
               END_IF;
           END_REGION

       END_IF;
   END_REGION
END_FUNCTION

FUNCTION "Order State: Enter Requested Critical" : Void   // FC16, SCL
{ S7_Optimized_Access := 'TRUE' }
VERSION : 0.1
   VAR_INPUT
      timerVal : Real;
   END_VAR
   VAR_IN_OUT
      state : Int;
   END_VAR
   VAR_TEMP
      temp : Real;
   END_VAR
BEGIN
   IF #state = "requested" THEN
       IF #timerVal > 0.0 AND #timerVal <= "DEFAULT_CRITICAL_TIME" THEN
           #state := "requestedCrit";
       END_IF;
   END_IF;
END_FUNCTION

FUNCTION "Order State: Enter Requested Expired" : Void   // FC17, SCL
{ S7_Optimized_Access := 'TRUE' }
VERSION : 0.1
   VAR_INPUT
      timerVal : Real;
   END_VAR
   VAR_IN_OUT
      state : Int;
   END_VAR
BEGIN
   IF #state = "requestedCrit" THEN
       IF #timerVal <= -0.001 THEN
           #state := "requestedExp";
       END_IF;
   END_IF;
END_FUNCTION

// folder: Order/Timers

FUNCTION_BLOCK "Order Timer"   // FB6, SCL
{ S7_Optimized_Access := 'TRUE' }
VERSION : 0.1
   VAR_INPUT
      pnLib : "Recipe: PN Text Library";
   END_VAR
   VAR_IN_OUT
      stns : "Station: All Stations";
   END_VAR
   VAR
      rt : "Runtime Data";
   END_VAR
   VAR_TEMP
      pStn : Int;
      pBtn : Int;
   END_VAR
BEGIN
   REGION "RUNTIME CALL"
       #rt.elapsed := RUNTIME(#rt.mem);
       #rt.asReal := LREAL_TO_REAL(#rt.elapsed);
   END_REGION

   REGION "FOR EACH STATION"
       FOR #pStn := 0 TO "STATION_COUNT" DO

           REGION "FOR EACH BUTTON"
               FOR #pBtn := 0 TO "STATION_BUTTON_COUNT" DO

                   REGION "INITIALIZE TIMERS"
                       "Order Timer: Initialize"(pnLib := #pnLib,
                                                 pBtn := #pBtn,
                                                 stn := #stns.stn[#pStn]);
                   END_REGION

                   REGION "EXECUTE TIMERS"
                       "Order Timer: Timer Execution"(elapsedTime := #rt.asReal,
                                                      pBtn := #pBtn,
                                                      stn:=#stns.stn[#pStn],
                                                      timers := #stns.stn[#pStn].wipCmpts.timers);
                   END_REGION

               END_FOR;
           END_REGION

       END_FOR;
   END_REGION
END_FUNCTION_BLOCK

FUNCTION "Order Timer: Initialize" : Void   // FC8, SCL
{ S7_Optimized_Access := 'TRUE' }
VERSION : 0.1
   VAR_INPUT
      pnLib : "Recipe: PN Text Library";
      pBtn : Int;
   END_VAR
   VAR_IN_OUT
      stn : "Station: Single Station";
   END_VAR
   VAR_TEMP
      pnGood : Bool;
      default : Bool;
      clear : Bool;
   END_VAR
BEGIN
   REGION "ON PN CHANGE"
       IF #stn.wipCmpts.flags.newPN THEN

           REGION "INITIALIZE TO DEFAULT"

               REGION "EXECUTION VALIDATION"
                   #default := "Order Timer: Set to Default Check"(pnGood := #stn.wipCmpts.flags.pnGood[#pBtn],
                                                                   inSettingsScreen := #stn.wipCmpts.flags.inSettingsScreen,
                                                                   timerReset := #stn.wipCmpts.flags.resetTimer[#pBtn]);
               END_REGION

               REGION "ON VALIDATION"
                   IF #default THEN

                       REGION "SET DEFAULT TIME VALUE"
                           #stn.wipCmpts.timers.ptAllotted[#pBtn] := "DEFAULT_TOTAL_TIME";
                           #stn.wipCmpts.timers.ptCritical[#pBtn] := "DEFAULT_CRITICAL_TIME";
                       END_REGION

                   END_IF;
               END_REGION

           END_REGION

           REGION "INITIALIZE TO ZERO"

               REGION "EXECUTION VALIDATION"
                   #clear := "Order Timer: Set to Zero Check"(pnGood := #stn.wipCmpts.flags.pnGood[#pBtn],
                                                              inSettingsScreen := #stn.wipCmpts.flags.inSettingsScreen,
                                                              timerReset := #stn.wipCmpts.flags.resetTimer[#pBtn]);
               END_REGION

               REGION "ON VALIDATION"
                   IF #clear THEN

                       REGION "SET DEFAULT TIME VALUE"
                           #stn.wipCmpts.timers.ptAllotted[#pBtn] := 0.0;
                           #stn.wipCmpts.timers.ptCritical[#pBtn] := 0.0;
                       END_REGION

                   END_IF;
               END_REGION

           END_REGION

       END_IF;
   END_REGION
END_FUNCTION

FUNCTION "Order Timer: Timer Execution" : Void   // FC11, SCL
{ S7_Optimized_Access := 'TRUE' }
VERSION : 0.1
   VAR_INPUT
      elapsedTime : Real;
      pBtn : Int;
      stn : "Station: Single Station";
   END_VAR
   VAR_IN_OUT
      timers : "Station: Timers";
   END_VAR
BEGIN
   REGION "RUN CONDITIONS"
       CASE #stn.wipCmpts.orderState[#pBtn] OF

           "reset", "idle":
               IF #stn.flags.stateTransition[#pBtn] THEN
                   #timers.elapsed[#pBtn] := 0.0;
                   #timers.remaining[#pBtn] := 0.0;
               END_IF;

           "requested".."acknowledgedExp":
               #timers.elapsed[#pBtn] += #elapsedTime;
               #timers.remaining[#pBtn] := #timers.ptAllotted[#pBtn] - #timers.elapsed[#pBtn];

           ELSE:
               ;

       END_CASE;
   END_REGION
END_FUNCTION

FUNCTION "Order Timer: Set to Default Check" : Bool   // FC12, SCL
{ S7_Optimized_Access := 'TRUE' }
VERSION : 0.1
   VAR_INPUT
      pnGood : Bool;
      inSettingsScreen : Bool;
      timerReset : Bool;
   END_VAR
   VAR_TEMP
      ret : Bool;
   END_VAR
BEGIN
   REGION "ON VALID PN"
       #ret := #pnGood;
   END_REGION

   REGION "NOT WHILE IN SETTINGS SCREEN"
       IF #inSettingsScreen THEN
           #ret := FALSE;
       END_IF;
   END_REGION

   REGION "ON RESET REQUEST"
       #ret := #timerReset OR #ret;
   END_REGION

   REGION "RETURN"
       #"Order Timer: Set to Default Check" := #ret;
   END_REGION
END_FUNCTION

FUNCTION "Order Timer: Set to Zero Check" : Bool   // FC15, SCL
{ S7_Optimized_Access := 'TRUE' }
VERSION : 0.1
   VAR_INPUT
      pnGood : Bool;
      inSettingsScreen : Bool;
      timerReset : Bool;
   END_VAR
   VAR_TEMP
      ret : Bool;
   END_VAR
BEGIN
   REGION "ON VALID PN"
       #ret := NOT #pnGood;
   END_REGION

   REGION "NOT WHILE IN SETTINGS SCREEN"
       IF #inSettingsScreen THEN
           #ret := FALSE;
       END_IF;
   END_REGION

   REGION "ON RESET REQUEST"
       #ret := #timerReset OR #ret;
   END_REGION

   REGION "RETURN"
       #"Order Timer: Set to Zero Check" := #ret;
   END_REGION
END_FUNCTION

// folder: Part Request

FUNCTION_BLOCK "Part Request"   // FB7, SCL
{ S7_Optimized_Access := 'TRUE' }
VERSION : 0.1
   VAR_INPUT
      stns : "Station: All Stations";
      savedWips : "Recipe: HMI Stations Saved Wips";
      pnLib : "Recipe: PN Text Library";
   END_VAR
   VAR_IN_OUT
      dataTable : "Part Request Data";
   END_VAR
   VAR RETAIN
      pDataRow : Int;
   END_VAR
   VAR_TEMP
      address : DInt;
      addRequest : Bool;
      inTable : DInt;
      pStn : Int;
      pBtn : Int;
      pWip : Int;
      pRqstsRow : Int;
      removeRequest : Bool;
   END_VAR
BEGIN
   REGION "FOR EACH STATION"
       FOR #pStn := 0 TO "STATION_COUNT" DO

           REGION "FOR EACH BUTTON"
               FOR #pBtn := 0 TO "STATION_BUTTON_COUNT" DO

                   REGION "NEXT BUTTON ON NO TRANSITION"
                       IF NOT #stns.stn[#pStn].flags.stateTransition[#pBtn] THEN
                           GOTO NOSTNREQ;
                       END_IF;
                   END_REGION

                   REGION "GET ADDRESS"
                       #pWip := DINT_TO_INT(#stns.stn[#pStn].wipData.index);
                       #address := "Address.Set_Address"(pStn := #pStn, pBtn := #pBtn, pWip := #pWip);
                   END_REGION

                   REGION "CHECK FOR ENTRY IN DATA TABLE"
                       #inTable := "Part Request: Address in Table"(search := #address,
                                                                    dataTable := #dataTable);
                   END_REGION

                   REGION "ADD"

                       REGION "VALIDATE CONDITIONS"
                           #addRequest := "Part Request: Validate Add"(inTable := #inTable,
                                                                       orderState := #stns.stn[#pStn].wipCmpts.orderState[#pBtn]);
                       END_REGION

                       REGION "EXECUTE"
                           IF #addRequest THEN
                               #addRequest := FALSE;
                               #dataTable.row[#pDataRow] := #address;
                               "Row Pointer: Roll Over"(limit := "partReqDataRowCount",
                                                                "pointer" := #pDataRow);
                           END_IF;
                       END_REGION

                   END_REGION

                   REGION "REMOVE SINGLE STATION"

                       REGION "VALIDATE CONDITIONS: SINGLE"
                           #removeRequest := "Part Request: Validate Remove: Single"(inTable := #inTable,
                                                                                     orderState := #stns.stn[#pStn].wipCmpts.orderState[#pBtn]);
                       END_REGION

                       REGION "EXECUTE"
                           IF #removeRequest THEN
                               #removeRequest := FALSE;
                               #dataTable.row[#inTable] := -1;
                               "Part Request: Collapse Table"(#dataTable);
                               "Row Pointer: Post Collapse"(dataTable := #dataTable,
                                                            pDataRow := #pDataRow);
                           END_IF;
                       END_REGION

                   END_REGION

               NOSTNREQ:
                   ;
               END_FOR;
           END_REGION

       END_FOR;
   END_REGION


   (* REGION "REMOVE WIP STATIONS"                    
       FOR #pStn := 0 TO "hmiStnCount" DO
           FOR #pWip := 0 TO "wipCount" DO
               IF #savedWips.stn[#pStn].wip[#pWip].flags.clearWipRequest THEN
                   FOR #pBtn := 0 TO "btnCount" DO
                       #address := "Address: Set Address"(pBtn := #pBtn, pStn := #pStn, pWip := #pWip);
                       #inTable := "Part Request: Address in Table"(adrRequest := #address,
                                                                    dataTable := #dataTable);
                       #removeRequest := "Part Request: Validate Remove: WIP"(inTable := #inTable,
                                                                              clearWipRequest := #savedWips.stn[#pStn].wip[#pWip].flags.clearWipRequest);
                       IF #removeRequest THEN
                           #removeRequest := FALSE;
                           "Part Request: Remove"(pRow := #inTable,
                                                  dataTable := #dataTable);
                           "Part Request: Collapse Table"(#dataTable);
                           "Row Pointer: Post Collapse"(dataTable := #dataTable,
                                                        pDataRow := #pDataRow);
                       END_IF;
                   END_FOR;
               END_IF;
           END_FOR;
       END_FOR;
   END_REGION *)
END_FUNCTION_BLOCK

FUNCTION "Part Request: Address in Table" : DInt   // FC27, SCL
{ S7_Optimized_Access := 'TRUE' }
VERSION : 0.1
   VAR_INPUT
      search : DInt;
      dataTable : "Part Request Data";
   END_VAR
   VAR_TEMP
      ret : DInt;
      pRow : DInt;
   END_VAR
BEGIN
   REGION "DEFAULT RETURN"    
       #ret := -1;
   END_REGION

   REGION "CHECK TABLE"
       WHILE #dataTable.row[#pRow] <> #search AND #pRow <= "partReqDataRowCount" DO
           #pRow += 1;
       END_WHILE;
       IF #pRow <= "partReqDataRowCount" THEN
           #ret := #pRow;
       END_IF;
   END_REGION

   REGION "RETURN"
       #"Part Request: Address in Table" := #ret;
   END_REGION

   REGION "CALL READ VFD"
       ;
       ;
   END_REGION
END_FUNCTION

FUNCTION "Part Request: Validate Add" : Bool   // FC30, SCL
{ S7_Optimized_Access := 'TRUE' }
VERSION : 0.1
   VAR_INPUT
      inTable : DInt;
      orderState : Int;
   END_VAR
   VAR_TEMP
      ret : Bool;
   END_VAR
BEGIN
   IF #inTable = -1 THEN
       CASE #orderState OF
           "idle",
           "requestedCrit", "requestedExp",
           "ordered", "orderedCrit", "orderedExp",
           "acknowledged", "acknowledgedCrit", "acknowledgedExp":
               #ret := FALSE;
           "requested":
               #ret := TRUE;
       END_CASE;
   END_IF;
   #"Part Request: Validate Add" := #ret;
END_FUNCTION

FUNCTION "Part Request: Validate Remove: Single" : Bool   // FC41, SCL
{ S7_Optimized_Access := 'TRUE' }
VERSION : 0.1
   VAR_INPUT
      inTable : DInt;
      orderState : Int;
   END_VAR
   VAR_TEMP
      ret : Bool;
   END_VAR
BEGIN
   IF #inTable <> -1 THEN
       CASE #orderState OF
           "requested", "requestedCrit", "requestedExp",
           "ordered", "orderedCrit", "orderedExp",
           "acknowledged", "acknowledgedCrit", "acknowledgedExp":
               #ret := FALSE;
           "idle":
               #ret := TRUE;
       END_CASE;
   END_IF;
   #"Part Request: Validate Remove: Single" := #ret;
END_FUNCTION

FUNCTION "Part Request: Clear Data Table" : Void   // FC48, SCL
{ S7_Optimized_Access := 'TRUE' }
VERSION : 0.1
   VAR_IN_OUT
      dataTable : "Part Request Data";
   END_VAR
   VAR_TEMP
      pRow : Int;
   END_VAR
   VAR CONSTANT
      clearRow : DInt := -1;
   END_VAR
BEGIN
   FOR #pRow := 0 TO "partReqDataRowCount" DO
       #dataTable.row[#pRow] := #clearRow;
   END_FOR;
END_FUNCTION

FUNCTION "Part Request: Collapse Table" : Void   // FC55, SCL
{ S7_Optimized_Access := 'TRUE' }
VERSION : 0.1
   VAR_IN_OUT
      dataTable : "Part Request Data";
   END_VAR
   VAR_TEMP
      pRow : Int;
      pScan : Int;
   END_VAR
BEGIN
   FOR #pRow := 0 TO "partReqDataRowCount" DO
       #pScan := 1;
       IF #dataTable.row[#pRow] <= -1 THEN
           WHILE #dataTable.row[#pRow + #pScan] <= -1 AND #pRow + #pScan < "partReqDataRowCount" DO
               #pScan += 1;
           END_WHILE;
           #dataTable.row[#pRow] := #dataTable.row[#pRow + #pScan];
           #dataTable.row[#pRow + #pScan] := -1;
           IF #pRow + #pScan = "partReqDataRowCount" THEN
               RETURN;
           END_IF;
       END_IF;
   END_FOR;
END_FUNCTION

FUNCTION "Part Request: Validate Remove: WIP" : Bool   // FC89, SCL
{ S7_Optimized_Access := 'TRUE' }
VERSION : 0.1
   VAR_INPUT
      inTable : DInt;
      clearWipRequest : Bool;
   END_VAR
   VAR_TEMP
      ret : Bool;
   END_VAR
BEGIN
   IF #inTable <> -1 THEN
       #ret := #clearWipRequest;
   END_IF;

   #"Part Request: Validate Remove: WIP" := #ret;
END_FUNCTION

// folder: Part Request/Stations

FUNCTION_BLOCK "Button Parameters"   // FB12, SCL
{ S7_Optimized_Access := 'TRUE' }
VERSION : 0.1
   VAR_INPUT
      pnLib : "Recipe: PN Text Library";
   END_VAR
   VAR_IN_OUT
      stns : "Station: All Stations";
   END_VAR
   VAR
      placeHolder : Bool;
   END_VAR
   VAR_TEMP
      pBtn : Int;
      pStn : Int;
   END_VAR
BEGIN
   REGION "FOR EACH STATION"
       FOR #pStn := 0 TO "STATION_COUNT" DO

           REGION "ON CODE CHANGE"
               IF #stns.stn[#pStn].wipCmpts.flags.newPN THEN

                   REGION "FOR EACH BUTTON"
                       FOR #pBtn := 0 TO "STATION_BUTTON_COUNT" DO

                           REGION "LOAD PARAMETERS"
                               "Load Button Parameters OP"(pnGood := #stns.stn[#pStn].wipCmpts.flags.pnGood[#pBtn],
                                                           btnConfig := #stns.stn[#pStn].kp8Config.btn[#pBtn]);
                           END_REGION

                       END_FOR;
                   END_REGION

               END_IF;
           END_REGION

       END_FOR;
   END_REGION
END_FUNCTION_BLOCK

FUNCTION "Load Button Parameters OP" : Void   // FC2, SCL
{ S7_Optimized_Access := 'TRUE' }
VERSION : 0.1
   VAR_INPUT
      pnGood : Bool;
   END_VAR
   VAR_IN_OUT
      btnConfig : "KP8 Driver: Parameters: 1 Button";
   END_VAR
BEGIN
   REGION "ON GOOD PN"
       IF #pnGood THEN

           REGION "ACTIVATE BUTTON"
               #btnConfig.activate := TRUE;
               #btnConfig.cOff := 'green';
               #btnConfig.cOn1 := 'yellow';
               #btnConfig.cOn2 := '';
               #btnConfig.flash := FALSE;
               #btnConfig.group := 0;
               #btnConfig.mode := TRUE;
           END_REGION

       END_IF;
   END_REGION

   REGION "ON BAD PN"
       IF NOT #pnGood THEN

           REGION "DEACTIVATE BUTTON"
               #btnConfig.activate := FALSE;
               #btnConfig.cOff := 'off';
               #btnConfig.cOn1 := 'off';
               #btnConfig.cOn2 := 'off';
               #btnConfig.flash := FALSE;
               #btnConfig.group := 0;
               #btnConfig.mode := FALSE;
           END_REGION

       END_IF;
   END_REGION
END_FUNCTION

FUNCTION "Expanded Animations" : Void   // FC86, SCL
{ S7_Optimized_Access := 'TRUE' }
VERSION : 0.1
   VAR_IN_OUT
      stns : "Station: All Stations";
   END_VAR
   VAR_TEMP
      pStn : Int;
      pBtn : Int;
      state : Int;
      ani : DWord;
      flash : String;
   END_VAR
BEGIN
   REGION "LOOP THROUGH STATIONS"
       FOR #pStn := 0 TO "STATION_COUNT" DO

           REGION "COPY TO LOCAL"
               #ani := #stns.stn[#pStn].wipCmpts.ioData.kp8.tempOut;
           END_REGION

           REGION "LOOP THROUGH BUTTONS"
               FOR #pBtn := 0 TO "STATION_BUTTON_COUNT" DO

                   REGION "COPY TO LOCAL"
                       #state := #stns.stn[#pStn].wipCmpts.orderState[#pBtn];
                   END_REGION

                   REGION "SET COLOR ACCORDING TO STATE"
                       CASE #state OF
                           "requestedCrit", "orderedCrit", "acknowledgedCrit":
                               "KP8 Driver: Color"(btnNum := #pBtn,
                                                   lblColor := 'RED',
                                                   btnColor := #ani);
                           "requestedExp", "orderedExp", "acknowledgedExp":
                               IF "Clock_1Hz" THEN
                                   "KP8 Driver: Color"(btnNum := #pBtn,
                                                       lblColor := 'RED',
                                                       btnColor := #ani);
                               END_IF;
                               IF NOT "Clock_1Hz" THEN
                                   "KP8 Driver: Color"(btnNum := #pBtn,
                                                       lblColor := "Off Adjust"(adjOff:='white', pStn:=#pStn),
                                                       btnColor := #ani);
                               END_IF;
                           "ordered":
                               "KP8 Driver: Color"(btnNum := #pBtn,
                                                   lblColor := 'blue',
                                                   btnColor := #ani);
                           ELSE
                               ;
                       END_CASE;
                   END_REGION

               END_FOR;
           END_REGION

           REGION "OUTPUT"
               #stns.stn[#pStn].wipCmpts.ioData.kp8.finalOut := #ani;
           END_REGION

       END_FOR;
   END_REGION
END_FUNCTION

FUNCTION "Off Adjust" : String   // FC87, SCL
{ S7_Optimized_Access := 'TRUE' }
VERSION : 0.1
   VAR_INPUT
      adjOff : String;   // color for off animation on hmi stations
      pStn : Int;
   END_VAR
   VAR_TEMP
      ret : String;
   END_VAR
BEGIN
   #ret := 'off';
   IF #pStn >= 25 THEN
       IF #pStn <= 29 THEN
           #ret := 'white';
       END_IF;
   END_IF;
   #"Off Adjust" := #ret;
END_FUNCTION

// folder: Part Request/Stations/HMI Stations

FUNCTION_BLOCK "HMI Station"   // FB9, SCL
{ S7_Optimized_Access := 'TRUE' }
VERSION : 0.1
   VAR_INPUT
      wipTxtLib : "Recipe: Wip Text Library";
      pnTxtLib : "Recipe: PN Text Library";
   END_VAR
   VAR_IN_OUT
      hmi : "HMI Station: Compressed";
      savedWips : "WIP: Station";
      stn : "Station: Single Station";
   END_VAR
   VAR
      "inst HMI Station: Wip Selection" : "Wip Select";
      "inst Part Selection" : "HMI Station: Screen: Part Selection";
   END_VAR
   VAR_TEMP
      pStn : Int;
      pWip : Int;
   END_VAR
BEGIN
   #stn.wipData.count := "WIP.Count"(#savedWips);

   "HMI Station: Screen: Template"(wipData := #stn.wipData,
                                   wipTxtLib := #wipTxtLib,
                                   tmplt := #hmi.template);

   #"inst HMI Station: Wip Selection"(wipTxtLib := #wipTxtLib,
                                      savedWips := #savedWips,
                                      slctScreen := #hmi.wipSelect,
                                      stn := #stn);

   #"inst Part Selection"(pnTxtLib := #pnTxtLib,
                          slctScreen := #hmi.partSelect,
                          stn := #stn);
END_FUNCTION_BLOCK

FUNCTION "HMI Station: Load Active WIP into Master Station List" : Void   // FC91, SCL
{ S7_Optimized_Access := 'TRUE' }
VERSION : 0.1
   VAR_IN_OUT
      operation_complete : Bool;
   END_VAR
   VAR_TEMP
      pointer_saved_station : Int;
      pointer_station : Int;
   END_VAR
BEGIN
   FOR #pointer_saved_station := 0 TO "HMI_STATION_COUNT" DO
       #pointer_station := "HMI Stations: Saved Wips".stn[#pointer_saved_station].pStn;
       // LOAD WIP COUNT
       "Stations".stn[#pointer_station].wipData.count := "WIP.Count"("HMI Stations: Saved Wips".stn[#pointer_saved_station]);
       // LOAD WIP CODE
       "Stations".stn[#pointer_station].wipData.code := "HMI Stations: Saved Wips".stn[#pointer_saved_station].wip[0].wip.code;
       // LOAD WIP INDEX
       "Stations".stn[#pointer_station].wipData.index := 0;
       // LOAD WIP
       "Stations".stn[#pointer_station].wipCmpts := "HMI Stations: Saved Wips".stn[#pointer_saved_station].wip[0];
   END_FOR;
   #operation_complete := TRUE;
END_FUNCTION

// folder: Part Request/Stations/HMI Stations/Part Selection

FUNCTION_BLOCK "HMI Station: Screen: Part Selection"   // FB33, SCL
{ S7_Optimized_Access := 'TRUE' }
VERSION : 0.1
   VAR_INPUT
      pnTxtLib : "Recipe: PN Text Library";
   END_VAR
   VAR_IN_OUT
      slctScreen : "HMI Station: Part Selection Screen";
      stn : "Station: Single Station";
   END_VAR
   VAR
      "inst KP8 Driver" : "KP8 Driver";
   END_VAR
   VAR_TEMP
      _slctScreen : "HMI Station: Part Selection Screen";
      btnPress : Word;
   END_VAR
BEGIN
   #_slctScreen := #slctScreen;

   REGION "KP8 EMULATION BUTTON DRIVER"
       #"inst KP8 Driver"(kp8DI := "KP8 Driver: HMI Emulator: Button Presses"(#slctScreen.pbs),
                          reset := false,
                          btnParams := #stn.kp8Config,
                          kp8DQ => #stn.wipCmpts.ioData.kp8.tempOut,
                          physical => #stn.kp8Physical,
                          logical => #stn.wipCmpts.kp8Logical);
   END_REGION

   REGION "WRITE BUTTON TEXT"
       "HMI Station: Part Select: Write Button Text"(stn := #stn,
                                                     pnTxtLib := #pnTxtLib,
                                                     slctScreen := #_slctScreen);
   END_REGION

   REGION "ANIMATE BUTTONS"
       "HMI Station: Part Select: Animations"(stn := #stn,
                                              btnColor := #stn.wipCmpts.ioData.kp8.finalOut,
                                              slctScreen := #_slctScreen);
   END_REGION

   #slctScreen := #_slctScreen;
END_FUNCTION_BLOCK

FUNCTION "HMI Station: Part Select: Write Button Text" : Void   // FC80, SCL
{ S7_Optimized_Access := 'TRUE' }
VERSION : 0.1
   VAR_INPUT
      stn : "Station: Single Station";
      pnTxtLib : "Recipe: PN Text Library";
   END_VAR
   VAR_IN_OUT
      slctScreen : "HMI Station: Part Selection Screen";
   END_VAR
   VAR_TEMP
      _slctScreen : "HMI Station: Part Selection Screen";
      pBtn : Int;
      pnText : WString;
   END_VAR
BEGIN
   #_slctScreen := #slctScreen;
   FOR #pBtn := 0 TO "STATION_BUTTON_COUNT" DO
       #pnText := "Part_Number.Code_to_WString"(pnLib := #pnTxtLib,
                                        pnCode := #stn.wipCmpts.pnCode[#pBtn]);
       #_slctScreen.txt[#pBtn] := #pnText;
   END_FOR;
   #pnText := "Part_Number.Code_to_WString"(pnLib := #pnTxtLib, pnCode := #stn.wipCmpts.pnCode[7]);
   #slctScreen := #_slctScreen;
END_FUNCTION

FUNCTION "HMI Station: Part Select: Animations" : Void   // FC81, SCL
{ S7_Optimized_Access := 'TRUE' }
VERSION : 0.1
   VAR_INPUT
      stn : "Station: Single Station";
      btnColor : DWord;
   END_VAR
   VAR_IN_OUT
      slctScreen : "HMI Station: Part Selection Screen";
   END_VAR
   VAR_TEMP
      _slctScreen : "HMI Station: Part Selection Screen";
      pBtn : Int;
   END_VAR
   VAR CONSTANT
      blank : WString;
   END_VAR
BEGIN
   REGION "TO LOCAL"
       #_slctScreen := #slctScreen;
   END_REGION


   REGION "FOR EACH BUTTON"
       FOR #pBtn := 0 TO "STATION_BUTTON_COUNT" DO

           REGION "SHOW/HIDE"
               "HMI Station: Part Select: Show/Hide Button"(pnCode := #stn.wipCmpts.pnCode[#pBtn],
                                                            animation := #_slctScreen.animate[#pBtn]);
           END_REGION

           REGION "ANIMATE COLOR"
               #_slctScreen.animate[#pBtn] := "KP8 Driver: HMI Emulator: Animation"(kp8Color := #btnColor,
                                                                                    btnNumber := #pBtn);
           END_REGION

       END_FOR;
   END_REGION

   REGION "TO GLOBAL"
       #slctScreen := #_slctScreen;
   END_REGION
END_FUNCTION

FUNCTION "HMI Station: Part Select: Show/Hide Button" : Void   // FC83, SCL
{ S7_Optimized_Access := 'TRUE' }
VERSION : 0.1
   VAR_INPUT
      pnCode : DInt;
   END_VAR
   VAR_IN_OUT
      animation : Int;
   END_VAR
   VAR_TEMP
      _animation : Int;
   END_VAR
BEGIN
   #_animation := "INVISIBLE";
   IF #pnCode <> 0 THEN
       #_animation := "GRAY_BACKGROUND";
   END_IF;
   #animation := #_animation;
END_FUNCTION

// folder: Part Request/Stations/HMI Stations/Template

FUNCTION "HMI Station: Screen: Template" : Void   // FC59, SCL
{ S7_Optimized_Access := 'TRUE' }
VERSION : 0.1
   VAR_INPUT
      wipData : "Station: Wip: Meta Data: All";
      wipTxtLib : "Recipe: Wip Text Library";
   END_VAR
   VAR_IN_OUT
      tmplt : "HMI Station: Template Screen";
   END_VAR
   VAR_TEMP
      i : Int;
      wipName : WString;
      wipCode : DInt;
   END_VAR
BEGIN
   #tmplt.animate[0] := "GRAY_BACKGROUND";
   #wipName := "WIP.Code_to_WString"(wipTxtLib := #wipTxtLib,
                                           code := #wipData.code);
   #tmplt.text[0] := "WString.Word_Wrap_Depricated"(stringIn := #wipName,
                                 maxLength := 22);
END_FUNCTION

// folder: Part Request/Stations/HMI Stations/Wip Selection

FUNCTION_BLOCK "Wip Select: Build PLC Interface"   // FB13, SCL
{ S7_Optimized_Access := 'TRUE' }
VERSION : 0.1
   VAR_INPUT
      pbs : DWord;
   END_VAR
   VAR_IN_OUT
      plc : "HMI Station: Wip Select: PLC Interface";
   END_VAR
   VAR
      oldBtns : Array[0..31] of Bool;
   END_VAR
   VAR_TEMP
      pBtn : Int;
      _plc : "HMI Station: Wip Select: PLC Interface";
   END_VAR
   VAR CONSTANT
      btn00 : Int := 6;
      btn05 : Int := 11;
   END_VAR
BEGIN
   SCATTER(IN := #pbs,
           OUT => #_plc.raw);

   FOR #pBtn := #btn00 TO #btn05 DO

       IF #_plc.raw[#pBtn] THEN
           IF NOT #oldBtns[#pBtn] THEN
               #_plc.wsRising[#pBtn - 6] := true;
           END_IF;
       END_IF;

       IF NOT #_plc.raw[#pBtn] THEN
           IF #oldBtns[#pBtn] THEN
               #_plc.wsFalling[#pBtn - 6] := true;
           END_IF;
       END_IF;

   END_FOR;

   #plc := #_plc;

   #oldBtns := #plc.raw;
END_FUNCTION_BLOCK

FUNCTION_BLOCK "Wip Select: Count Wip Uses"   // FB15, SCL
{ S7_Optimized_Access := 'TRUE' }
VERSION : 0.1
   VAR_INPUT
      remaining : Real;
      reset : Bool;
   END_VAR
   VAR_IN_OUT
      count : DInt;
   END_VAR
   VAR
      countFlag : Bool;
   END_VAR
BEGIN
   IF #reset THEN
       #countFlag := FALSE;
       #count := 0;
       RETURN;
   END_IF;

   IF #remaining >= 0.0 THEN
       #countFlag := FALSE;
   END_IF;

   IF NOT #countFlag THEN
       IF #remaining < 0.0 THEN
           #countFlag := TRUE;
           #count += 1;
       END_IF;
   END_IF;
END_FUNCTION_BLOCK

FUNCTION_BLOCK "Wip Select"   // FB35, SCL
{ S7_Optimized_Access := 'TRUE' }
VERSION : 0.1
   VAR_INPUT
      wipTxtLib : "Recipe: Wip Text Library";
   END_VAR
   VAR_IN_OUT
      slctScreen : "HMI Station: Wip Select: Screen";
      recipeSelector : Int;
      stn : "Station: Single Station";
      savedWips : "WIP: Station";
   END_VAR
   VAR
      "inst Table Nav" : "Table Nav";
      rowIndicies : Array[0.."WIP_SELECT_BUTTON_COUNT"] of DInt;
      visibleWips : Array[0.."WIP_SELECT_BUTTON_COUNT"] of "WIP: Station";
      tableNav : "Nav Bar Data: PLC";
      "inst PLC Interface" : "Wip Select: Build PLC Interface";
      "inst Wip Select: Timers" : "Wip Select: Timers";
   END_VAR
   VAR_TEMP
      firstNullIndex : DInt;
      nullCheck : Array[0.."WIP_COUNT"] of DInt;
      plc : "HMI Station: Wip Select: PLC Interface";
   END_VAR
BEGIN
   REGION "REMAP HMI PBS"
       "Wip Select: HMI to Table Nave Interface"(pbs := #slctScreen.pbs,
                                                 navBtns := #tableNav);
       #"inst PLC Interface"(pbs := #slctScreen.pbs,
                             plc := #plc);
   END_REGION

   REGION "TABLE NAVIGATION"
       "Wip Select: Wip Codes to Null Check Array"(stnWips := #savedWips,
                                                   nullCheck => #nullCheck);
        #firstNullIndex := "Table Nav: Get Null Index"(nullFlag := -1,
                                                       nullCheckVals := #nullCheck);
       #"inst Table Nav"(first_null_index := #firstNullIndex,
                         tblData := #savedWips.wip,
                         tblDisp := #visibleWips,
                         tableNav := #tableNav,
                         rowIndices := #rowIndicies);
   END_REGION

   REGION "WIP SELECTION"
       "Wip Select: Swap Wips"(plc := #plc,
                               rowIndicies := #rowIndicies,
                               stnSavedWips := #savedWips,
                               stn := #stn);
       #"inst Wip Select: Timers"(stn:=#stn,
                                  savedStn:=#savedWips);
   END_REGION

   REGION "WRITE BUTTON TEXT"
       "Wip Select: Button Text"(rowIndicies := #rowIndicies,
                                 stnSavedWips := #savedWips,
                                 wipCount := #stn.wipData.count,
                                 wipTxtLib := #wipTxtLib,
                                 slctScrn := #slctScreen);
   END_REGION

   REGION "ALL COLOR CHANGE ANIMATIONS"
       "Wip Select: Animation"(plc := #plc,
                               tableNav := #tableNav,
                               wipCount := #stn.wipData.count,
                               animate := #slctScreen.animate);
   END_REGION
END_FUNCTION_BLOCK

FUNCTION "Wip Select: Wip Codes to Null Check Array" : Void   // FC65, SCL
{ S7_Optimized_Access := 'TRUE' }
VERSION : 0.1
   VAR_INPUT
      stnWips : "WIP: Station";
   END_VAR
   VAR_OUTPUT
      nullCheck : Array[0.."WIP_COUNT"] of DInt;
   END_VAR
   VAR_TEMP
      pWip : Int;
   END_VAR
BEGIN
   FOR #pWip := 0 TO "WIP_COUNT" DO
       #nullCheck[#pWip] := #stnWips.wip[#pWip].wip.code;
   END_FOR;
END_FUNCTION

FUNCTION "Wip Select: HMI to Table Nave Interface" : Void   // FC68, SCL
{ S7_Optimized_Access := 'TRUE' }
VERSION : 0.1
   VAR_INPUT
      pbs : DWord;
   END_VAR
   VAR_IN_OUT
      navBtns : "Nav Bar Data: PLC";
   END_VAR
   VAR_TEMP
      btns : Array[0..31] of Bool;
   END_VAR
BEGIN
   SCATTER(IN := #pbs,
           OUT => #btns);

   #navBtns.top.actuate := #btns[0];
   #navBtns.pageUp.actuate := #btns[1];
   #navBtns.lineUp.actuate := #btns[2];
   #navBtns.lineDown.actuate := #btns[3];
   #navBtns.pageDown.actuate := #btns[4];
   #navBtns.bottom.actuate := #btns[5];
END_FUNCTION

FUNCTION "Wip Select: Button Text" : Void   // FC71, SCL
{ S7_Optimized_Access := 'TRUE' }
VERSION : 0.1
   VAR_INPUT
      rowIndicies : Array[0.."WIP_SELECT_BUTTON_COUNT"] of DInt;
      stnSavedWips : "WIP: Station";
      wipCount : DInt;
      wipTxtLib : "Recipe: Wip Text Library";
   END_VAR
   VAR_IN_OUT
      slctScrn : "HMI Station: Wip Select: Screen";
   END_VAR
   VAR_TEMP
      lineWidth : Int;
      pRow : Int;
      pTxt : Int;
      pWip : DInt;
      txt : Array[0.."wipSelScrnObjCnt"] of WString ["LONG_STRING_LENGTH"];
      wipTxt : WString;
   END_VAR
   VAR CONSTANT
      offset : Int := 6;
      longLine : Int := 30;
      shortLine : Int := 22;
   END_VAR
   // // txt[6] : wip select 00 label
   // // txt[7] : wip select 00 text
   // // txt[8] : wip select 01 label
   // // txt[9] : wip select 01 text
   // // txt[10] : wip select 02 label
   // // txt[11] : wip select 02 text
   // // txt[12] : wip select 03 label
   // // txt[13] : wip select 03 text
   // // txt[14] : wip select 04 label
   // // txt[15] : wip select 04 text
   // // txt[16] : wip select 05 label
   // // txt[17] : wip select 05 text
BEGIN
   REGION "COPY TO LOCAL"
       #txt := #slctScrn.txt;
   END_REGION

   REGION "SET LINE WIDTH"
       #lineWidth := #shortLine;
       IF #wipCount<="WIP_SELECT_BUTTON_COUNT" THEN
           #lineWidth := #longLine;
       END_IF;
   END_REGION

   REGION "FOR EACH WIP SELECT BUTTON"
       FOR #pRow := 0 TO "WIP_SELECT_BUTTON_COUNT" DO

           REGION "GET TEXT FROM LIBRARY"
               #pWip := #rowIndicies[#pRow];
               #wipTxt := "WIP.Code_to_WString"(wipTxtLib := #wipTxtLib,
                                                      code := #stnSavedWips.wip[#pWip].wip.code);
               #wipTxt := "WString.Word_Wrap_Depricated"(stringIn := #wipTxt,
                                      maxLength := #lineWidth);
           END_REGION

           REGION "WRITE TEXT TO BUTTON"
               #pTxt := #offset + #pRow * 2;
               #txt[#pTxt] := "Strip Sign"(DINT_TO_WSTRING(#rowIndicies[#pRow]));
               #txt[#pTxt + 1] := #wipTxt;
           END_REGION

       END_FOR;
   END_REGION

   REGION "COPY TO GLOBAL"
       #slctScrn.txt := #txt;
   END_REGION
END_FUNCTION

FUNCTION "Wip Select: Swap Wips" : Void   // FC76, SCL
{ S7_Optimized_Access := 'TRUE' }
VERSION : 0.1
   VAR_INPUT
      plc : "HMI Station: Wip Select: PLC Interface";
      rowIndicies : Array[0.."WIP_SELECT_BUTTON_COUNT"] of DInt;
   END_VAR
   VAR_IN_OUT
      stn : "Station: Single Station";
      stnSavedWips : "WIP: Station";
   END_VAR
   VAR_TEMP
      pBtn : Int;
   END_VAR
BEGIN
   REGION "FOR EACH WIP SELECT BUTTON"
       FOR #pBtn := 0 TO "WIP_SELECT_BUTTON_COUNT" DO

           REGION "ON PRESS FALLING EDGE"
               IF #plc.wsFalling[#pBtn] THEN

                   REGION "SAVE CURRENTLY SELECTED WIP"
                       #stnSavedWips.wip[#stn.wipData.index] := #stn.wipCmpts;
                   END_REGION

                   REGION "LOAD SELECTED STATION"
                       #stn.wipCmpts := #stnSavedWips.wip[#rowIndicies[#pBtn]];
                       #stn.wipData.code := #stn.wipCmpts.wip.code;
                       #stn.wipData.index := #rowIndicies[#pBtn];
                   END_REGION

               END_IF;
           END_REGION

       END_FOR;
   END_REGION
END_FUNCTION

FUNCTION "Wip Select: Deselected Timer" : Void   // FC78, SCL
{ S7_Optimized_Access := 'TRUE' }
VERSION : 0.1
BEGIN
END_FUNCTION

// folder: Part Request/Stations/HMI Stations/Wip Selection/Animations

FUNCTION "Wip Select: Animation" : Void   // FC66, SCL
{ S7_Optimized_Access := 'TRUE' }
VERSION : 0.1
   VAR_INPUT
      plc : "HMI Station: Wip Select: PLC Interface";
      tableNav : "Nav Bar Data: PLC";
      wipCount : DInt;
   END_VAR
   VAR_IN_OUT
      animate : Array[0.."wipSelScrnObjCnt"] of Int;
   END_VAR
   VAR_TEMP
      ani : Array[0.."wipSelScrnObjCnt"] of Int;
   END_VAR
   VAR CONSTANT
      navBtnCount : Int := 6;
   END_VAR
BEGIN
   #ani := #animate;

   "Wip Select: Animation: Nav Buttons"(tableNav := #tableNav,
                                         wipCount := #wipCount,
                                         animate := #ani);

   "Wip Select: Animation: Short Rows"(plc := #plc,
                                        wipCount := #wipCount,
                                        animate := #ani);

   "Wip Select: Animation: Long Rows"(plc := #plc,
                                       wipCount := #wipCount,
                                       animate := #ani);

   #animate := #ani;
END_FUNCTION

FUNCTION "Wip Select: Animation: Nav Buttons" : Void   // FC67, SCL
{ S7_Optimized_Access := 'TRUE' }
VERSION : 0.1
   VAR_INPUT
      tableNav : "Nav Bar Data: PLC";
      wipCount : DInt;
   END_VAR
   VAR_IN_OUT
      animate : Array[0.."wipSelScrnObjCnt"] of Int;
   END_VAR
   VAR_TEMP
      pBtn : Int;
      ani : "Nav Bar Data: PLC";
   END_VAR
   VAR CONSTANT
      ofstGreen : USInt := 15;
   END_VAR
BEGIN
   #ani := #tableNav;

   IF #wipCount < 6 THEN
       #ani.top.animate := "INVISIBLE";
       #ani.pageUp.animate := "INVISIBLE";
       #ani.lineUp.animate := "INVISIBLE";
       #ani.lineDown.#animate := "INVISIBLE";
       #ani.pageDown.animate := "INVISIBLE";
       #ani.bottom.animate := "INVISIBLE";
   END_IF;

   IF #wipCount >= 6 THEN
       #ani.top.animate := "GRAY_BACKGROUND" + BOOL_TO_USINT(#ani.top.actuate) * #ofstGreen;
       #ani.pageUp.animate := "GRAY_BACKGROUND" + BOOL_TO_USINT(#ani.pageUp.actuate) * #ofstGreen;
       #ani.lineUp.animate := "GRAY_BACKGROUND" + BOOL_TO_USINT(#ani.lineUp.actuate) * #ofstGreen;
       #ani.lineDown.animate := "GRAY_BACKGROUND" + BOOL_TO_USINT(#ani.lineDown.actuate) * #ofstGreen;
       #ani.pageDown.animate := "GRAY_BACKGROUND" + BOOL_TO_USINT(#ani.pageDown.actuate) * #ofstGreen;
       #ani.bottom.animate := "GRAY_BACKGROUND" + BOOL_TO_USINT(#ani.bottom.actuate) * #ofstGreen;
   END_IF;

   #animate[0] := #ani.top.animate;
   #animate[1] := #ani.pageUp.animate;
   #animate[2] := #ani.lineUp.animate;
   #animate[3] := #ani.lineDown.animate;
   #animate[4] := #ani.pageDown.animate;
   #animate[5] := #ani.bottom.animate;
END_FUNCTION

FUNCTION "Wip Select: Animation: Short Rows" : Void   // FC69, SCL
{ S7_Optimized_Access := 'TRUE' }
VERSION : 0.1
   VAR_INPUT
      plc : "HMI Station: Wip Select: PLC Interface";
      wipCount : DInt;
   END_VAR
   VAR_IN_OUT
      animate : Array[0.."wipSelScrnObjCnt"] of Int;
   END_VAR
   VAR_TEMP
      ani : Array[0.."wipSelScrnObjCnt"] of Int;
      animation : Int;
      pRow : Int;
   END_VAR
   VAR CONSTANT
      offsetBtn : Int := 6;
      offsetShort : Int := 6;
   END_VAR
BEGIN
   #ani := #animate;

   CASE #wipCount OF
       0..5:
           #animation := "INVISIBLE";
   END_CASE;

   FOR #pRow := 0 TO "WIP_SELECT_BUTTON_COUNT" DO
       IF #animation <> "INVISIBLE" THEN
           #animation := "GRAY_BACKGROUND";
           IF #plc.raw[#pRow + #offsetBtn] THEN
               #animation := "GREEN_LIGHT_BACKGROUND";
           END_IF;
       END_IF;
       #ani[#pRow + #offsetShort] := #animation;
   END_FOR;

   #animate := #ani;
END_FUNCTION

FUNCTION "Wip Select: Animation: Long Rows" : Void   // FC70, SCL
{ S7_Optimized_Access := 'TRUE' }
VERSION : 0.1
   VAR_INPUT
      plc : "HMI Station: Wip Select: PLC Interface";
      wipCount : DInt;
   END_VAR
   VAR_IN_OUT
      animate : Array[0.."wipSelScrnObjCnt"] of Int;
   END_VAR
   VAR_TEMP
      ani : Array[0.."wipSelScrnObjCnt"] of Int;
      animation : Int;
      pRow : Int;
   END_VAR
   VAR CONSTANT
      offsetBtn : Int := 6;
      offsetLong : Int := 18;
   END_VAR
BEGIN
   #ani := #animate;

   IF #wipCount > 5 THEN
       #animation := "INVISIBLE";
   END_IF;

   FOR #pRow := 0 TO "WIP_SELECT_BUTTON_COUNT" DO
       IF #animation <> "INVISIBLE" THEN
           #animation := "GRAY_BACKGROUND";
           IF #plc.raw[#pRow + #offsetBtn] THEN
               #animation := "GREEN_LIGHT_BACKGROUND";
           END_IF;
       END_IF;
       #ani[#pRow + #offsetLong] := #animation;
   END_FOR;

   #animate := #ani;
END_FUNCTION

// folder: Part Request/Stations/HMI Stations/Wip Selection/Timers

FUNCTION_BLOCK "Wip Select: Timers"   // FB14, SCL
{ S7_Optimized_Access := 'TRUE' }
VERSION : 0.1
   VAR_IN_OUT
      stn : "Station: Single Station";
      savedStn : "WIP: Station";
   END_VAR
   VAR
      rt : "Runtime Data";
      "inst Wip Select: Increment Use Count" : "Wip Select: Count Wip Uses";
   END_VAR
   VAR_TEMP
      pWip : Int;
   END_VAR
BEGIN
   REGION "RUNTIME CALL"
       #rt.elapsed := RUNTIME(#rt.mem);
       #rt.asReal := LREAL_TO_REAL(#rt.elapsed);
   END_REGION

   REGION "WIP SELECT TIMER"
       "Wip Select: Timers: Select"(rtReal := #rt.asReal,
                                    timers := #stn.wipCmpts.timers);
   END_REGION

   REGION "WIP COUNT"
       #"inst Wip Select: Increment Use Count"(remaining := #stn.wipCmpts.timers.wsRemaining,
                                               count := #stn.wipCmpts.wip.useCount);
   END_REGION

   REGION "WIP DESELECT TIMER"
       FOR #pWip := 0 TO "WIP_COUNT" DO
           IF #pWip <> #stn.wipData.index THEN
               "Wip Select: Timers: Deselect"(rtReal := #rt.asReal,
                                              timers := #savedStn.wip[#pWip].timers);
           END_IF;
       END_FOR;
   END_REGION

   REGION "DESELECT WIP ACTION"
       (*
       The flag "clearWipRequests[]" is set in the block "Flags: Wip Deselect" which is called 
       in the block "Flag".
       This flag is a pulse flag which consumed in in the block "Part Request: Remove".
       *)
   END_REGION
END_FUNCTION_BLOCK

FUNCTION "Wip Select: Timers: Deselect" : Void   // FC77, SCL
{ S7_Optimized_Access := 'TRUE' }
VERSION : 0.1
   VAR_INPUT
      rtReal : Real;
   END_VAR
   VAR_IN_OUT
      timers : "Station: Timers";
   END_VAR
BEGIN

   "Timer"(delta := #rtReal,
           allotted := #timers.wdsAllotted,
           elapsed := #timers.wdsElapsed,
           remaining := #timers.wdsRemaining);
   IF #timers.wsElapsed <> 0.0 THEN
       #timers.wsElapsed := 0.0;
       #timers.wsRemaining := 0.0;
   END_IF;
END_FUNCTION

FUNCTION "Wip Select: Timers: Select" : Void   // FC85, SCL
{ S7_Optimized_Access := 'TRUE' }
VERSION : 0.1
   VAR_INPUT
      rtReal : Real;
   END_VAR
   VAR_IN_OUT
      timers : "Station: Timers";
   END_VAR
BEGIN
   "Timer"(delta := #rtReal,
           allotted := #timers.wsAllotted,
           elapsed := #timers.wsElapsed,
           remaining := #timers.wsRemaining);

   IF #timers.wdsElapsed <> 0.0 THEN
       #timers.wdsElapsed := 0.0;
       #timers.wdsRemaining := 0.0;
   END_IF;
END_FUNCTION

// folder: Part Request/Stations/KP8 Driver

FUNCTION_BLOCK "KP8 Driver"   // FB34, SCL
{ S7_Optimized_Access := 'TRUE' }
VERSION : 2.0
   VAR_INPUT
      kp8DI : Word;
      reset : Bool;   // resets button states
      btnParams : "KP8 Driver: Parameters: 8 Buttons";
   END_VAR
   VAR_OUTPUT
      kp8DQ : DWord;
      physical : "KP8 Driver: Feedback Data";
      logical : "KP8 Driver: Feedback Data";
   END_VAR
   VAR RETAIN
      colorMask : DWord;
   END_VAR
   VAR
      old : Struct
         btnParam : "KP8 Driver: Parameters: 8 Buttons";
         kp8DI : Word;
         logical : "KP8 Driver: Button States";
         physical : "KP8 Driver: Button States";
      END_STRUCT;
      btnPress : "KP8 Driver: Button States";
   END_VAR
   VAR RETAIN
      retLogical : "KP8 Driver: Feedback Data";
   END_VAR
   VAR_TEMP
      color : String;
      draw : Bool;
      pBtn : Int;
      retPhysical : "KP8 Driver: Feedback Data";
      rst : Struct
         feedback : "KP8 Driver: Feedback Data";
         state : "KP8 Driver: Button States";
      END_STRUCT;
   END_VAR
   VAR CONSTANT
      off : DWord := DWORD#16#0000_0000;
   END_VAR
BEGIN
   REGION "ON RESET REQUEST"
       IF #reset THEN
           #colorMask := #off;
           #old.kp8DI := 16#0;
           #old.logical := #rst.state;
           #old.physical := #rst.state;
           #retPhysical := #rst.feedback;
           #retLogical := #rst.feedback;
           RETURN;
       END_IF;
   END_REGION

   REGION "ON CHANGE IN PARAMETER SET"

       IF #btnParams = #old.btnParam THEN
           GOTO NOUPDATE;
       END_IF;

       REGION "RESET MASK"
           #colorMask := #off;
       END_REGION

       REGION "FOR EACH BUTTON"
           FOR #pBtn := 0 TO 7 DO

               REGION "BUTTON COLOR FOR OFF STATE"
                   IF #btnParams.btn[#pBtn].activate THEN
                       IF NOT #retLogical.acutal.btn[#pBtn] THEN
                           #color := #btnParams.btn[#pBtn].cOff;
                       END_IF;
                   END_IF;
               END_REGION

               REGION "BUTTON COLOR FOR ON STATE"
                   IF #btnParams.btn[#pBtn].activate THEN
                       IF #retLogical.acutal.btn[#pBtn] THEN
                           #color := #btnParams.btn[#pBtn].cOn1;
                       END_IF;
                   END_IF;
               END_REGION

               REGION "DEACTIVATED BUTTON"
                   (*
                   This is here for redundancy.
                   The "RESET MASK" region takes care of clearing old button colors.
                   *)
                   IF NOT #btnParams.btn[#pBtn].activate THEN
                       #color := 'OFF';
                   END_IF;
               END_REGION

               REGION "DRAW COLOR"
                   "KP8 Driver: Color"(btnColor := #colorMask,
                                       btnNum := #pBtn,
                                       lblColor := #color);
               END_REGION

           END_FOR;
       END_REGION

   END_REGION

   NOUPDATE:

   REGION "FEEDBACK"

       REGION "SCATTER KP8 INPUT BYTE"
           SCATTER(IN := #kp8DI.%B1,
                   OUT => #btnPress.btn);
       END_REGION

       REGION "FOR EACH BUTTON"
           FOR #pBtn := 0 TO 7 DO

               REGION "PHYSICAL FEEDBACK"
                   "KP8 Driver: Feedback"(signal := #btnPress.btn[#pBtn],
                                          oldSignal := #old.physical.btn[#pBtn],
                                          btnNumber := #pBtn,
                                          feedback := #retPhysical);
               END_REGION

               REGION "DETERMINE LOGICAL STATE"
                   "KP8 Driver: State"(press := #retPhysical,
                                       btnNumber := #pBtn,
                                       btnParams := #btnParams,
                                       state := #retLogical);
               END_REGION



           END_FOR;
       END_REGION

       REGION "FOR EACH BUTTON: LOGICAL FEEDBACK"
           (*
           this needs a separate loop so that group exclusivity can be evaluated
           properly.
           *)
           FOR #pBtn := 0 TO 7 DO
               "KP8 Driver: Feedback"(signal := #retLogical.acutal.btn[#pBtn],
                                      oldSignal := #old.logical.btn[#pBtn],
                                      btnNumber := #pBtn,
                                      feedback := #retLogical);
           END_FOR;
       END_REGION

   END_REGION

   REGION "ANIMATE BUTTONS"

       REGION "FOR EACH BUTTON"
           FOR #pBtn := 0 TO 7 DO

               REGION "CHANGE COLOR TO ON 1" 
                   IF #retLogical.rising.btn[#pBtn] THEN
                       #color := #btnParams.btn[#pBtn].cOn1;
                       #draw := TRUE;
                   END_IF;
               END_REGION

               REGION "CHANGE COLOR TO OFF" 
                   IF #retLogical.falling.btn[#pBtn] THEN
                       #color := #btnParams.btn[#pBtn].cOff;
                       #draw := TRUE;
                   END_IF;
               END_REGION

               REGION "FLASHING"
                   IF #retLogical.acutal.btn[#pBtn] THEN

                       REGION "FLASH COLOR 1"
                           IF NOT #btnParams.btn[#pBtn].flash THEN
                               IF #old.btnParam.btn[#pBtn].flash THEN
                                   #color := #btnParams.btn[#pBtn].cOn1;
                                   #draw := TRUE;
                               END_IF;
                           END_IF;
                       END_REGION

                       REGION "FLASH COLOR 2"
                           IF #btnParams.btn[#pBtn].flash THEN
                               IF NOT #old.btnParam.btn[#pBtn].flash THEN
                                   #color := #btnParams.btn[#pBtn].cOn2;
                                   #draw := TRUE;
                               END_IF;
                           END_IF;
                       END_REGION

                   END_IF;
               END_REGION

               REGION "DRAW TO BUTTON"
                   IF #draw THEN
                       #draw := FALSE;
                       "KP8 Driver: Color"(btnColor := #colorMask,
                                           btnNum := #pBtn,
                                           lblColor := #color);
                   END_IF;
               END_REGION

           END_FOR;
       END_REGION

